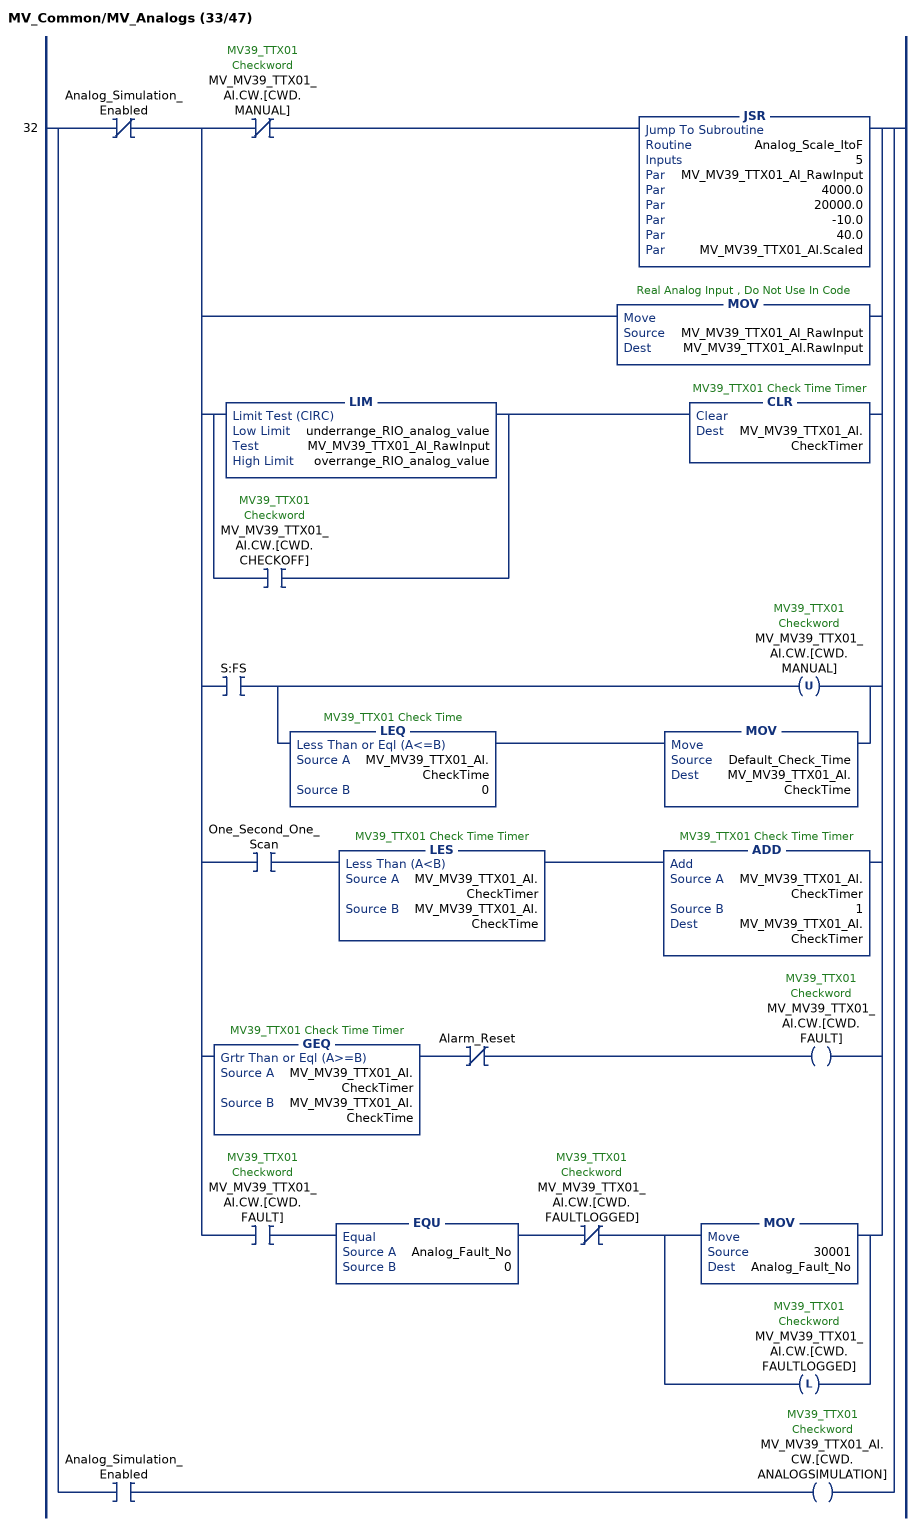
   32: [XIO(Analog_Simulation_Enabled) [XIO(MV_MV39_TTX01_AI.CW.[CWD.MANUAL]) JSR(Analog_Scale_ItoF,5,MV_MV39_TTX01_AI_RawInput,4000.0,20000.0,-10.0,40.0,MV_MV39_TTX01_AI.Scaled) ,MOV(MV_MV39_TTX01_AI_RawInput,MV_MV39_TTX01_AI.RawInput) ,[LIM(underrange_RIO_analog_value,MV_MV39_TTX01_AI_RawInput,overrange_RIO_analog_value) ,XIC(MV_MV39_TTX01_AI.CW.[CWD.CHECKOFF]) ] CLR(MV_MV39_TTX01_AI.CheckTimer) ,XIC(S:FS) [OTU(MV_MV39_TTX01_AI.CW.[CWD.MANUAL]) ,LEQ(MV_MV39_TTX01_AI.CheckTime,0) MOV(Default_Check_Time,MV_MV39_TTX01_AI.CheckTime) ] ,XIC(One_Second_One_Scan) LES(MV_MV39_TTX01_AI.CheckTimer,MV_MV39_TTX01_AI.CheckTime) ADD(MV_MV39_TTX01_AI.CheckTimer,1,MV_MV39_TTX01_AI.CheckTimer) ,GEQ(MV_MV39_TTX01_AI.CheckTimer,MV_MV39_TTX01_AI.CheckTime) XIO(Alarm_Reset) OTE(MV_MV39_TTX01_AI.CW.[CWD.FAULT]) ,XIC(MV_MV39_TTX01_AI.CW.[CWD.FAULT]) EQU(Analog_Fault_No,0) XIO(MV_MV39_TTX01_AI.CW.[CWD.FAULTLOGGED]) [MOV(30001,Analog_Fault_No) ,OTL(MV_MV39_TTX01_AI.CW.[CWD.FAULTLOGGED]) ] ] ,XIC(Analog_Simulation_Enabled) OTE(MV_MV39_TTX01_AI.CW.[CWD.ANALOGSIMULATION]) ];
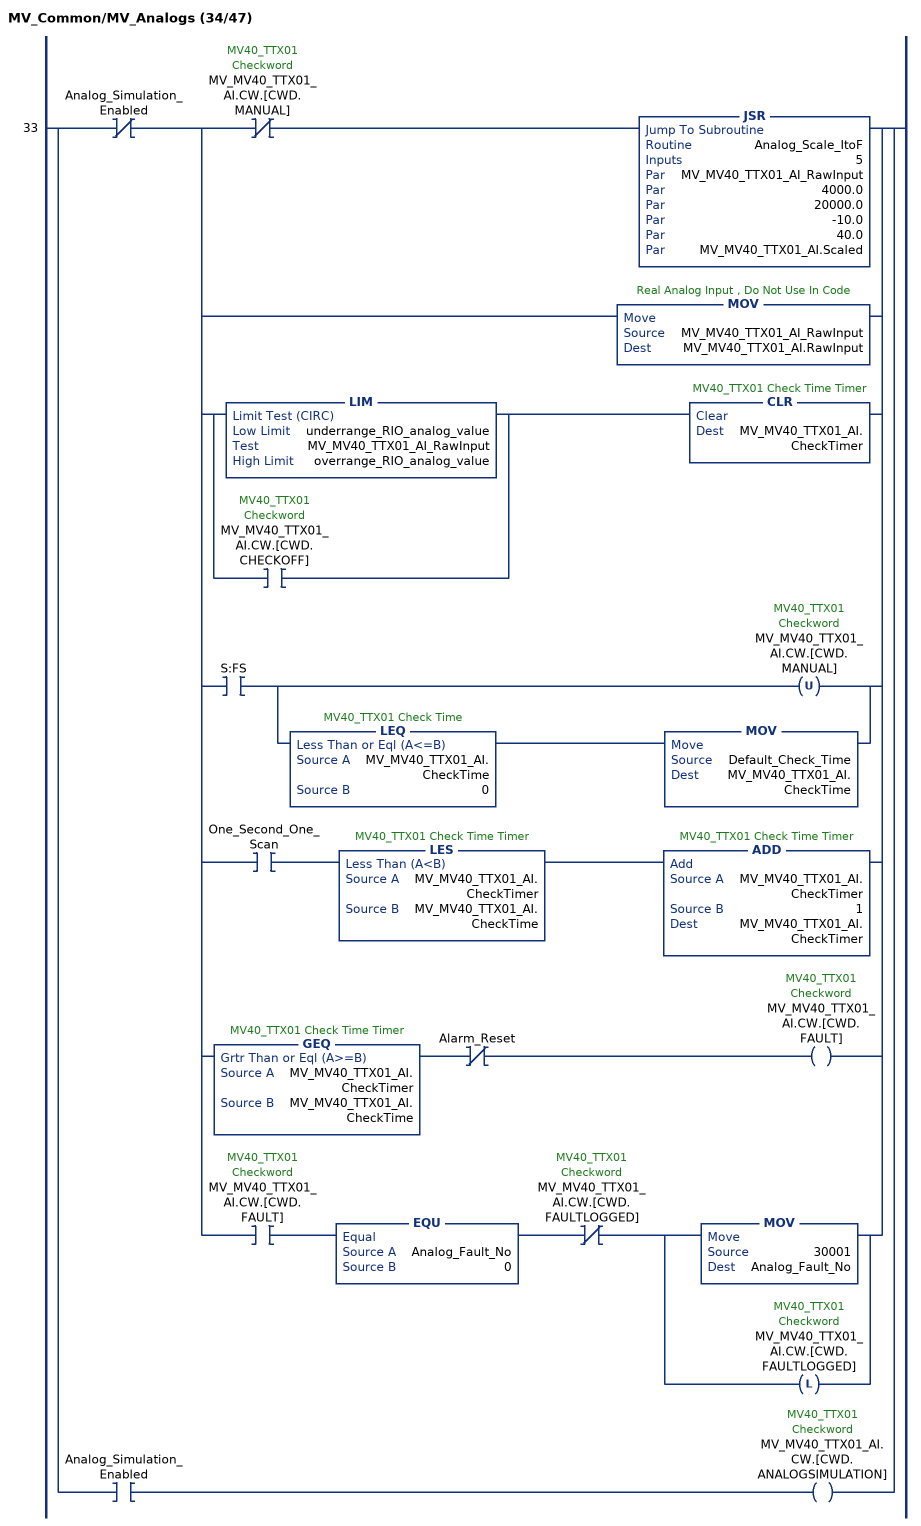
   33: [XIO(Analog_Simulation_Enabled) [XIO(MV_MV40_TTX01_AI.CW.[CWD.MANUAL]) JSR(Analog_Scale_ItoF,5,MV_MV40_TTX01_AI_RawInput,4000.0,20000.0,-10.0,40.0,MV_MV40_TTX01_AI.Scaled) ,MOV(MV_MV40_TTX01_AI_RawInput,MV_MV40_TTX01_AI.RawInput) ,[LIM(underrange_RIO_analog_value,MV_MV40_TTX01_AI_RawInput,overrange_RIO_analog_value) ,XIC(MV_MV40_TTX01_AI.CW.[CWD.CHECKOFF]) ] CLR(MV_MV40_TTX01_AI.CheckTimer) ,XIC(S:FS) [OTU(MV_MV40_TTX01_AI.CW.[CWD.MANUAL]) ,LEQ(MV_MV40_TTX01_AI.CheckTime,0) MOV(Default_Check_Time,MV_MV40_TTX01_AI.CheckTime) ] ,XIC(One_Second_One_Scan) LES(MV_MV40_TTX01_AI.CheckTimer,MV_MV40_TTX01_AI.CheckTime) ADD(MV_MV40_TTX01_AI.CheckTimer,1,MV_MV40_TTX01_AI.CheckTimer) ,GEQ(MV_MV40_TTX01_AI.CheckTimer,MV_MV40_TTX01_AI.CheckTime) XIO(Alarm_Reset) OTE(MV_MV40_TTX01_AI.CW.[CWD.FAULT]) ,XIC(MV_MV40_TTX01_AI.CW.[CWD.FAULT]) EQU(Analog_Fault_No,0) XIO(MV_MV40_TTX01_AI.CW.[CWD.FAULTLOGGED]) [MOV(30001,Analog_Fault_No) ,OTL(MV_MV40_TTX01_AI.CW.[CWD.FAULTLOGGED]) ] ] ,XIC(Analog_Simulation_Enabled) OTE(MV_MV40_TTX01_AI.CW.[CWD.ANALOGSIMULATION]) ];
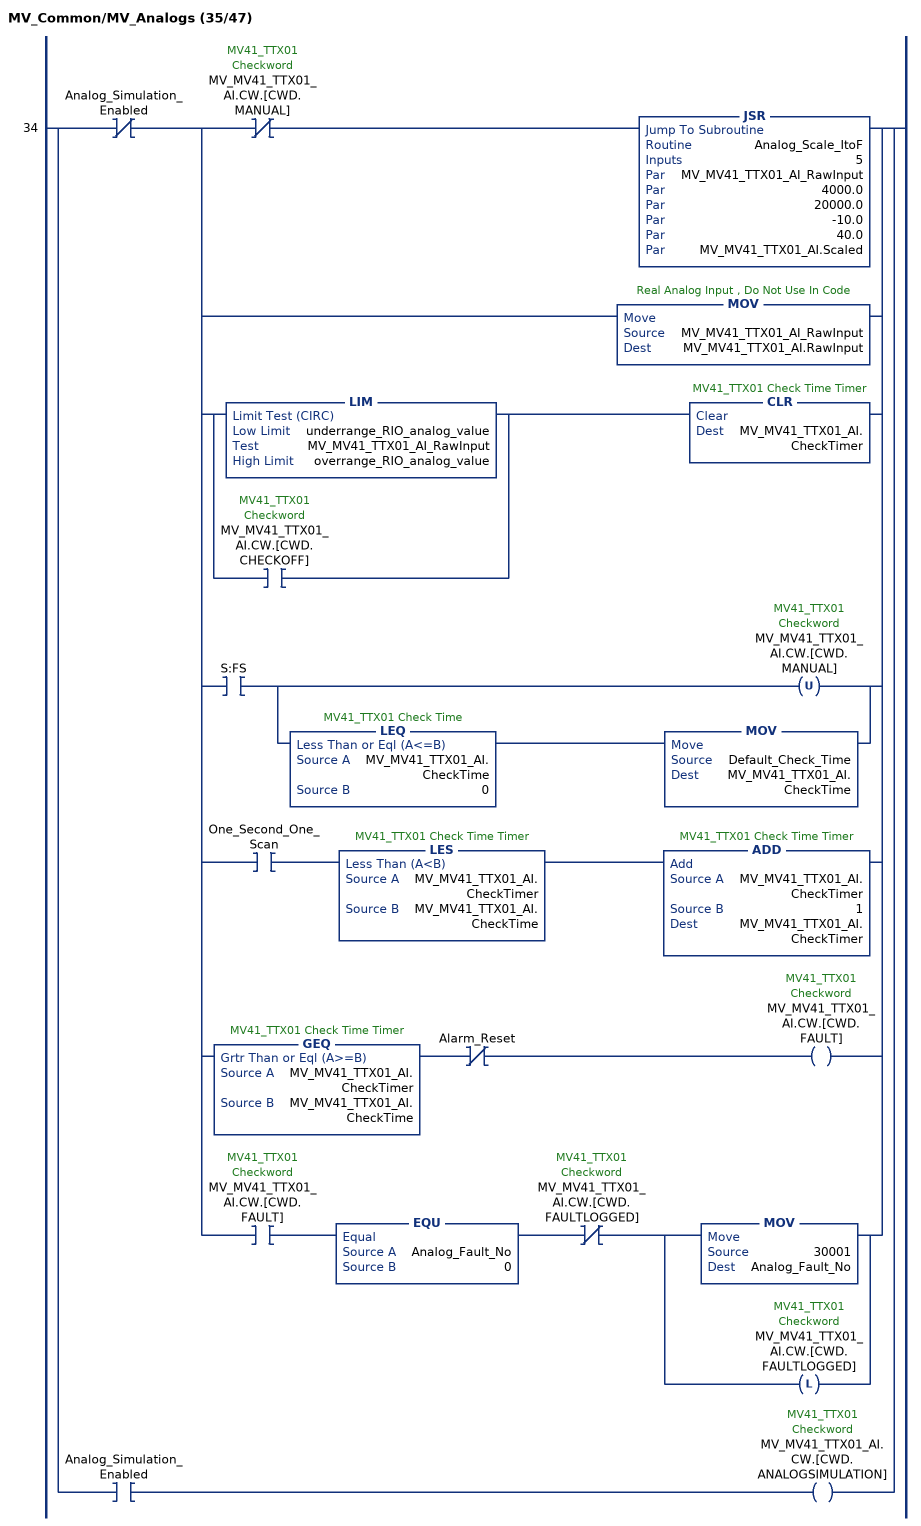
   34: [XIO(Analog_Simulation_Enabled) [XIO(MV_MV41_TTX01_AI.CW.[CWD.MANUAL]) JSR(Analog_Scale_ItoF,5,MV_MV41_TTX01_AI_RawInput,4000.0,20000.0,-10.0,40.0,MV_MV41_TTX01_AI.Scaled) ,MOV(MV_MV41_TTX01_AI_RawInput,MV_MV41_TTX01_AI.RawInput) ,[LIM(underrange_RIO_analog_value,MV_MV41_TTX01_AI_RawInput,overrange_RIO_analog_value) ,XIC(MV_MV41_TTX01_AI.CW.[CWD.CHECKOFF]) ] CLR(MV_MV41_TTX01_AI.CheckTimer) ,XIC(S:FS) [OTU(MV_MV41_TTX01_AI.CW.[CWD.MANUAL]) ,LEQ(MV_MV41_TTX01_AI.CheckTime,0) MOV(Default_Check_Time,MV_MV41_TTX01_AI.CheckTime) ] ,XIC(One_Second_One_Scan) LES(MV_MV41_TTX01_AI.CheckTimer,MV_MV41_TTX01_AI.CheckTime) ADD(MV_MV41_TTX01_AI.CheckTimer,1,MV_MV41_TTX01_AI.CheckTimer) ,GEQ(MV_MV41_TTX01_AI.CheckTimer,MV_MV41_TTX01_AI.CheckTime) XIO(Alarm_Reset) OTE(MV_MV41_TTX01_AI.CW.[CWD.FAULT]) ,XIC(MV_MV41_TTX01_AI.CW.[CWD.FAULT]) EQU(Analog_Fault_No,0) XIO(MV_MV41_TTX01_AI.CW.[CWD.FAULTLOGGED]) [MOV(30001,Analog_Fault_No) ,OTL(MV_MV41_TTX01_AI.CW.[CWD.FAULTLOGGED]) ] ] ,XIC(Analog_Simulation_Enabled) OTE(MV_MV41_TTX01_AI.CW.[CWD.ANALOGSIMULATION]) ];
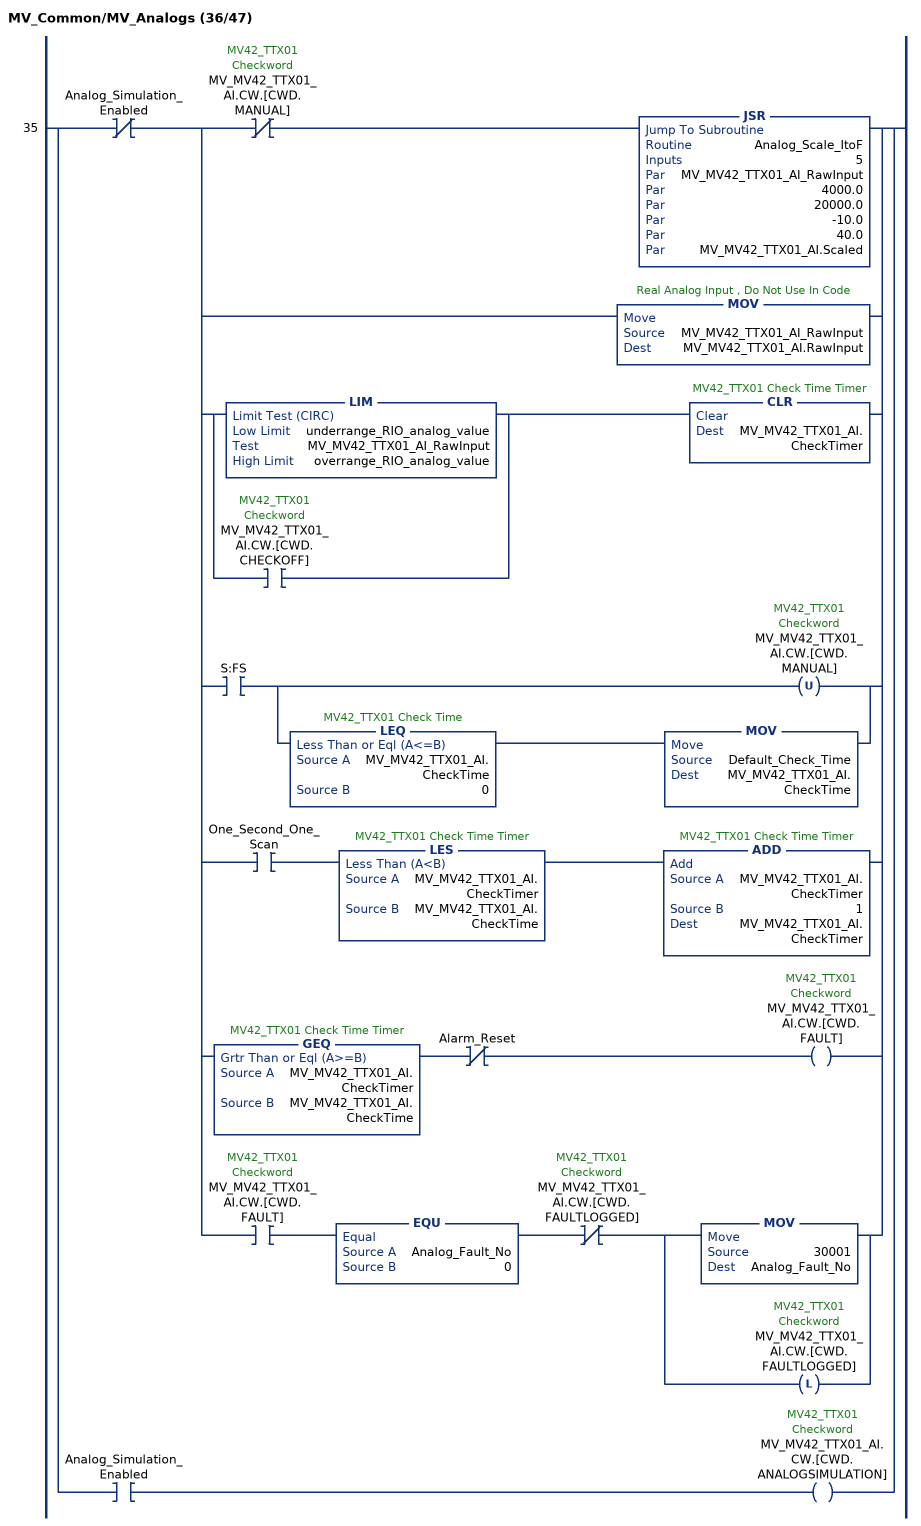
   35: [XIO(Analog_Simulation_Enabled) [XIO(MV_MV42_TTX01_AI.CW.[CWD.MANUAL]) JSR(Analog_Scale_ItoF,5,MV_MV42_TTX01_AI_RawInput,4000.0,20000.0,-10.0,40.0,MV_MV42_TTX01_AI.Scaled) ,MOV(MV_MV42_TTX01_AI_RawInput,MV_MV42_TTX01_AI.RawInput) ,[LIM(underrange_RIO_analog_value,MV_MV42_TTX01_AI_RawInput,overrange_RIO_analog_value) ,XIC(MV_MV42_TTX01_AI.CW.[CWD.CHECKOFF]) ] CLR(MV_MV42_TTX01_AI.CheckTimer) ,XIC(S:FS) [OTU(MV_MV42_TTX01_AI.CW.[CWD.MANUAL]) ,LEQ(MV_MV42_TTX01_AI.CheckTime,0) MOV(Default_Check_Time,MV_MV42_TTX01_AI.CheckTime) ] ,XIC(One_Second_One_Scan) LES(MV_MV42_TTX01_AI.CheckTimer,MV_MV42_TTX01_AI.CheckTime) ADD(MV_MV42_TTX01_AI.CheckTimer,1,MV_MV42_TTX01_AI.CheckTimer) ,GEQ(MV_MV42_TTX01_AI.CheckTimer,MV_MV42_TTX01_AI.CheckTime) XIO(Alarm_Reset) OTE(MV_MV42_TTX01_AI.CW.[CWD.FAULT]) ,XIC(MV_MV42_TTX01_AI.CW.[CWD.FAULT]) EQU(Analog_Fault_No,0) XIO(MV_MV42_TTX01_AI.CW.[CWD.FAULTLOGGED]) [MOV(30001,Analog_Fault_No) ,OTL(MV_MV42_TTX01_AI.CW.[CWD.FAULTLOGGED]) ] ] ,XIC(Analog_Simulation_Enabled) OTE(MV_MV42_TTX01_AI.CW.[CWD.ANALOGSIMULATION]) ];
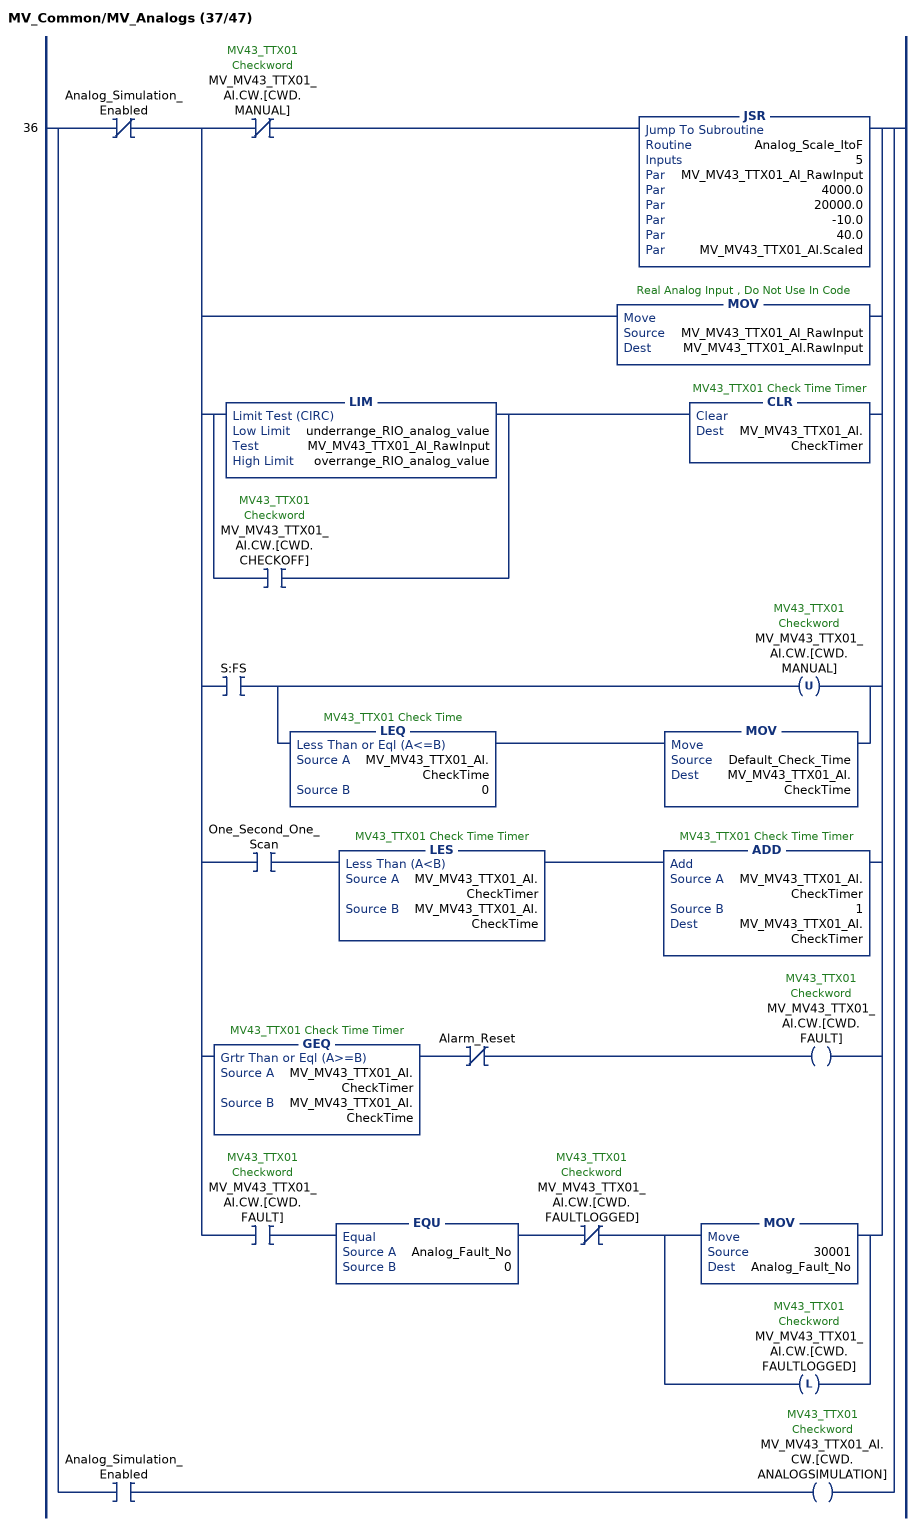
   36: [XIO(Analog_Simulation_Enabled) [XIO(MV_MV43_TTX01_AI.CW.[CWD.MANUAL]) JSR(Analog_Scale_ItoF,5,MV_MV43_TTX01_AI_RawInput,4000.0,20000.0,-10.0,40.0,MV_MV43_TTX01_AI.Scaled) ,MOV(MV_MV43_TTX01_AI_RawInput,MV_MV43_TTX01_AI.RawInput) ,[LIM(underrange_RIO_analog_value,MV_MV43_TTX01_AI_RawInput,overrange_RIO_analog_value) ,XIC(MV_MV43_TTX01_AI.CW.[CWD.CHECKOFF]) ] CLR(MV_MV43_TTX01_AI.CheckTimer) ,XIC(S:FS) [OTU(MV_MV43_TTX01_AI.CW.[CWD.MANUAL]) ,LEQ(MV_MV43_TTX01_AI.CheckTime,0) MOV(Default_Check_Time,MV_MV43_TTX01_AI.CheckTime) ] ,XIC(One_Second_One_Scan) LES(MV_MV43_TTX01_AI.CheckTimer,MV_MV43_TTX01_AI.CheckTime) ADD(MV_MV43_TTX01_AI.CheckTimer,1,MV_MV43_TTX01_AI.CheckTimer) ,GEQ(MV_MV43_TTX01_AI.CheckTimer,MV_MV43_TTX01_AI.CheckTime) XIO(Alarm_Reset) OTE(MV_MV43_TTX01_AI.CW.[CWD.FAULT]) ,XIC(MV_MV43_TTX01_AI.CW.[CWD.FAULT]) EQU(Analog_Fault_No,0) XIO(MV_MV43_TTX01_AI.CW.[CWD.FAULTLOGGED]) [MOV(30001,Analog_Fault_No) ,OTL(MV_MV43_TTX01_AI.CW.[CWD.FAULTLOGGED]) ] ] ,XIC(Analog_Simulation_Enabled) OTE(MV_MV43_TTX01_AI.CW.[CWD.ANALOGSIMULATION]) ];
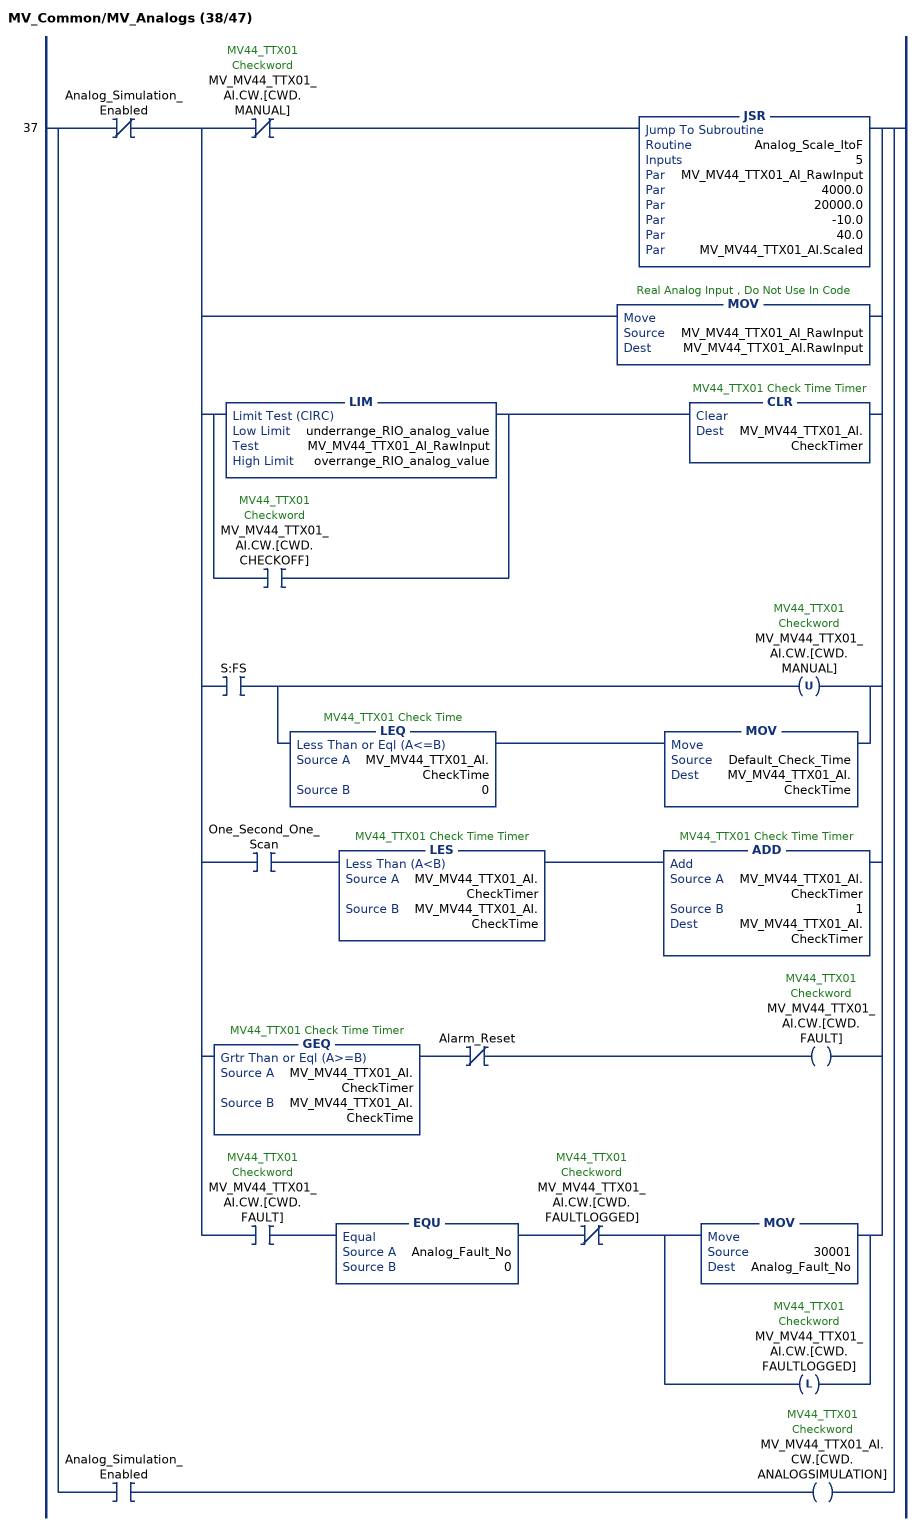
   37: [XIO(Analog_Simulation_Enabled) [XIO(MV_MV44_TTX01_AI.CW.[CWD.MANUAL]) JSR(Analog_Scale_ItoF,5,MV_MV44_TTX01_AI_RawInput,4000.0,20000.0,-10.0,40.0,MV_MV44_TTX01_AI.Scaled) ,MOV(MV_MV44_TTX01_AI_RawInput,MV_MV44_TTX01_AI.RawInput) ,[LIM(underrange_RIO_analog_value,MV_MV44_TTX01_AI_RawInput,overrange_RIO_analog_value) ,XIC(MV_MV44_TTX01_AI.CW.[CWD.CHECKOFF]) ] CLR(MV_MV44_TTX01_AI.CheckTimer) ,XIC(S:FS) [OTU(MV_MV44_TTX01_AI.CW.[CWD.MANUAL]) ,LEQ(MV_MV44_TTX01_AI.CheckTime,0) MOV(Default_Check_Time,MV_MV44_TTX01_AI.CheckTime) ] ,XIC(One_Second_One_Scan) LES(MV_MV44_TTX01_AI.CheckTimer,MV_MV44_TTX01_AI.CheckTime) ADD(MV_MV44_TTX01_AI.CheckTimer,1,MV_MV44_TTX01_AI.CheckTimer) ,GEQ(MV_MV44_TTX01_AI.CheckTimer,MV_MV44_TTX01_AI.CheckTime) XIO(Alarm_Reset) OTE(MV_MV44_TTX01_AI.CW.[CWD.FAULT]) ,XIC(MV_MV44_TTX01_AI.CW.[CWD.FAULT]) EQU(Analog_Fault_No,0) XIO(MV_MV44_TTX01_AI.CW.[CWD.FAULTLOGGED]) [MOV(30001,Analog_Fault_No) ,OTL(MV_MV44_TTX01_AI.CW.[CWD.FAULTLOGGED]) ] ] ,XIC(Analog_Simulation_Enabled) OTE(MV_MV44_TTX01_AI.CW.[CWD.ANALOGSIMULATION]) ];
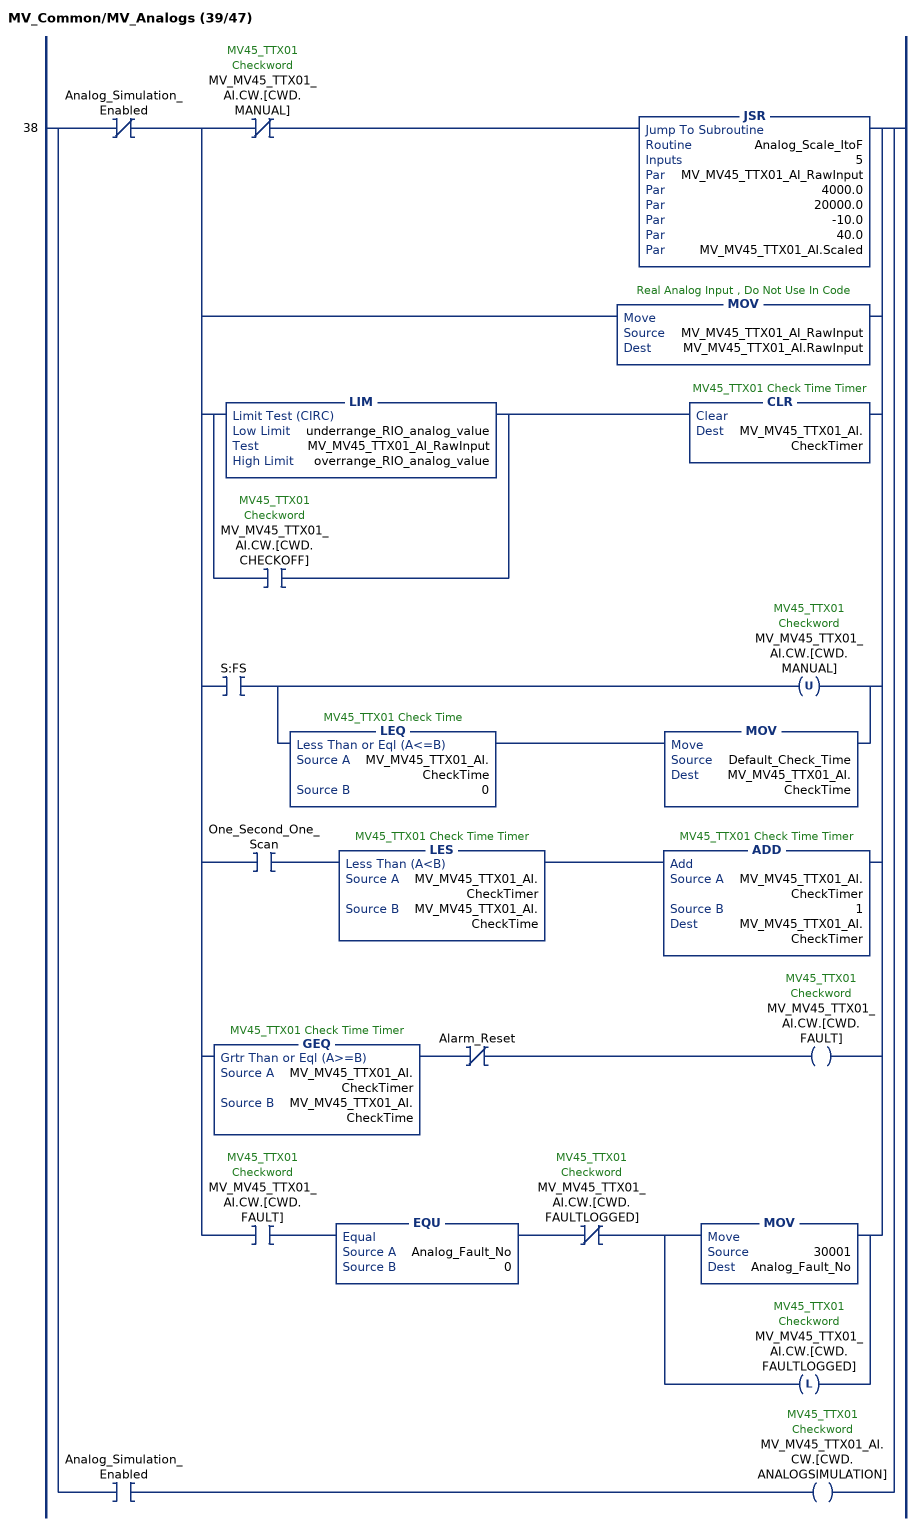
   38: [XIO(Analog_Simulation_Enabled) [XIO(MV_MV45_TTX01_AI.CW.[CWD.MANUAL]) JSR(Analog_Scale_ItoF,5,MV_MV45_TTX01_AI_RawInput,4000.0,20000.0,-10.0,40.0,MV_MV45_TTX01_AI.Scaled) ,MOV(MV_MV45_TTX01_AI_RawInput,MV_MV45_TTX01_AI.RawInput) ,[LIM(underrange_RIO_analog_value,MV_MV45_TTX01_AI_RawInput,overrange_RIO_analog_value) ,XIC(MV_MV45_TTX01_AI.CW.[CWD.CHECKOFF]) ] CLR(MV_MV45_TTX01_AI.CheckTimer) ,XIC(S:FS) [OTU(MV_MV45_TTX01_AI.CW.[CWD.MANUAL]) ,LEQ(MV_MV45_TTX01_AI.CheckTime,0) MOV(Default_Check_Time,MV_MV45_TTX01_AI.CheckTime) ] ,XIC(One_Second_One_Scan) LES(MV_MV45_TTX01_AI.CheckTimer,MV_MV45_TTX01_AI.CheckTime) ADD(MV_MV45_TTX01_AI.CheckTimer,1,MV_MV45_TTX01_AI.CheckTimer) ,GEQ(MV_MV45_TTX01_AI.CheckTimer,MV_MV45_TTX01_AI.CheckTime) XIO(Alarm_Reset) OTE(MV_MV45_TTX01_AI.CW.[CWD.FAULT]) ,XIC(MV_MV45_TTX01_AI.CW.[CWD.FAULT]) EQU(Analog_Fault_No,0) XIO(MV_MV45_TTX01_AI.CW.[CWD.FAULTLOGGED]) [MOV(30001,Analog_Fault_No) ,OTL(MV_MV45_TTX01_AI.CW.[CWD.FAULTLOGGED]) ] ] ,XIC(Analog_Simulation_Enabled) OTE(MV_MV45_TTX01_AI.CW.[CWD.ANALOGSIMULATION]) ];
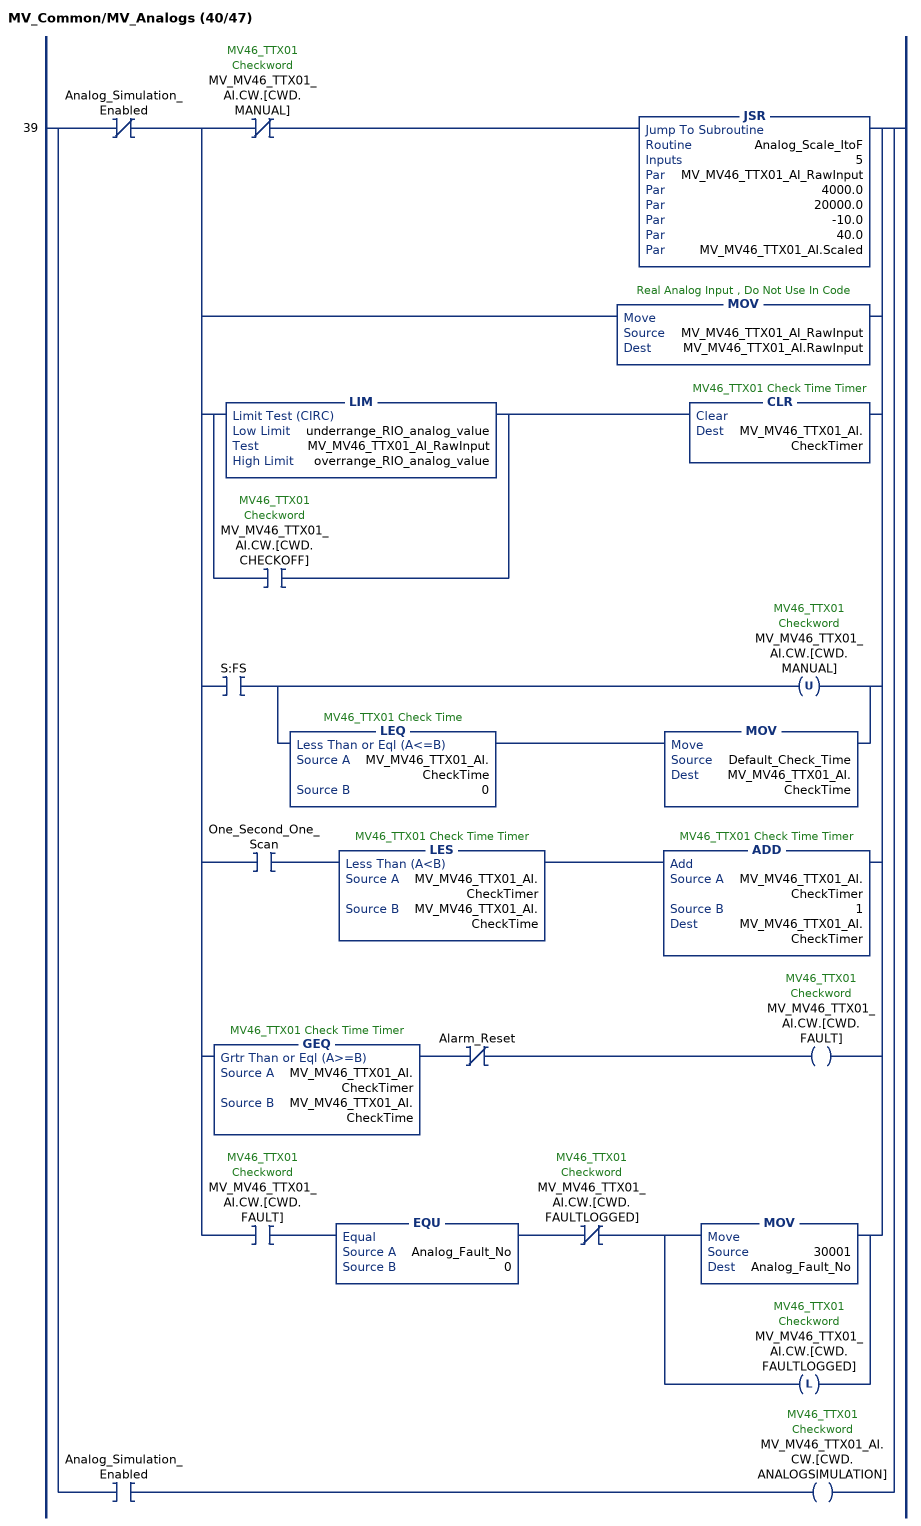
   39: [XIO(Analog_Simulation_Enabled) [XIO(MV_MV46_TTX01_AI.CW.[CWD.MANUAL]) JSR(Analog_Scale_ItoF,5,MV_MV46_TTX01_AI_RawInput,4000.0,20000.0,-10.0,40.0,MV_MV46_TTX01_AI.Scaled) ,MOV(MV_MV46_TTX01_AI_RawInput,MV_MV46_TTX01_AI.RawInput) ,[LIM(underrange_RIO_analog_value,MV_MV46_TTX01_AI_RawInput,overrange_RIO_analog_value) ,XIC(MV_MV46_TTX01_AI.CW.[CWD.CHECKOFF]) ] CLR(MV_MV46_TTX01_AI.CheckTimer) ,XIC(S:FS) [OTU(MV_MV46_TTX01_AI.CW.[CWD.MANUAL]) ,LEQ(MV_MV46_TTX01_AI.CheckTime,0) MOV(Default_Check_Time,MV_MV46_TTX01_AI.CheckTime) ] ,XIC(One_Second_One_Scan) LES(MV_MV46_TTX01_AI.CheckTimer,MV_MV46_TTX01_AI.CheckTime) ADD(MV_MV46_TTX01_AI.CheckTimer,1,MV_MV46_TTX01_AI.CheckTimer) ,GEQ(MV_MV46_TTX01_AI.CheckTimer,MV_MV46_TTX01_AI.CheckTime) XIO(Alarm_Reset) OTE(MV_MV46_TTX01_AI.CW.[CWD.FAULT]) ,XIC(MV_MV46_TTX01_AI.CW.[CWD.FAULT]) EQU(Analog_Fault_No,0) XIO(MV_MV46_TTX01_AI.CW.[CWD.FAULTLOGGED]) [MOV(30001,Analog_Fault_No) ,OTL(MV_MV46_TTX01_AI.CW.[CWD.FAULTLOGGED]) ] ] ,XIC(Analog_Simulation_Enabled) OTE(MV_MV46_TTX01_AI.CW.[CWD.ANALOGSIMULATION]) ];
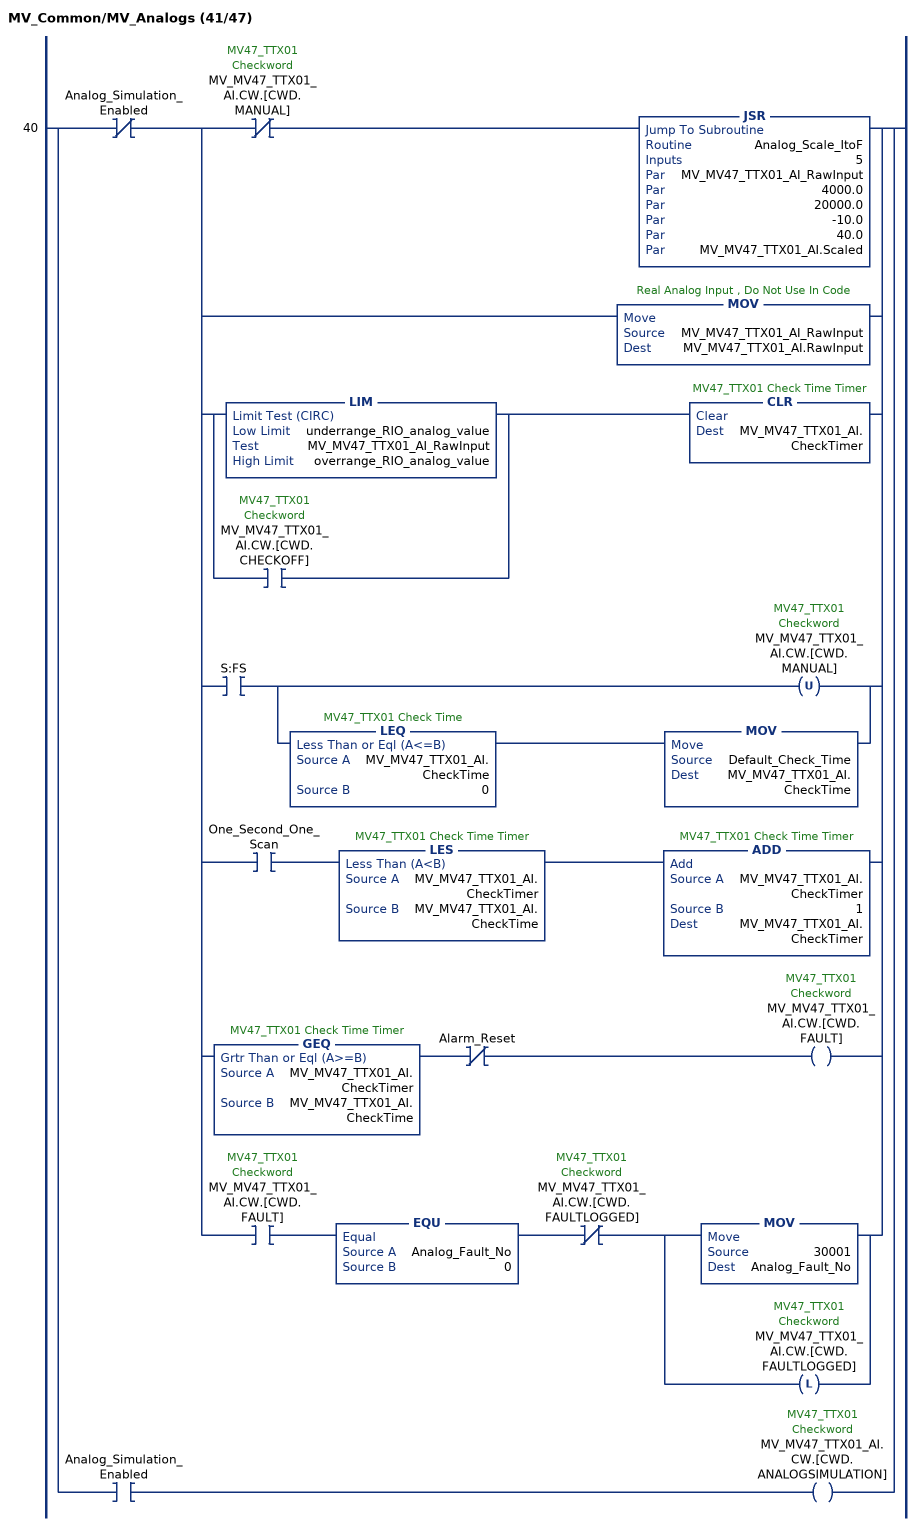
   40: [XIO(Analog_Simulation_Enabled) [XIO(MV_MV47_TTX01_AI.CW.[CWD.MANUAL]) JSR(Analog_Scale_ItoF,5,MV_MV47_TTX01_AI_RawInput,4000.0,20000.0,-10.0,40.0,MV_MV47_TTX01_AI.Scaled) ,MOV(MV_MV47_TTX01_AI_RawInput,MV_MV47_TTX01_AI.RawInput) ,[LIM(underrange_RIO_analog_value,MV_MV47_TTX01_AI_RawInput,overrange_RIO_analog_value) ,XIC(MV_MV47_TTX01_AI.CW.[CWD.CHECKOFF]) ] CLR(MV_MV47_TTX01_AI.CheckTimer) ,XIC(S:FS) [OTU(MV_MV47_TTX01_AI.CW.[CWD.MANUAL]) ,LEQ(MV_MV47_TTX01_AI.CheckTime,0) MOV(Default_Check_Time,MV_MV47_TTX01_AI.CheckTime) ] ,XIC(One_Second_One_Scan) LES(MV_MV47_TTX01_AI.CheckTimer,MV_MV47_TTX01_AI.CheckTime) ADD(MV_MV47_TTX01_AI.CheckTimer,1,MV_MV47_TTX01_AI.CheckTimer) ,GEQ(MV_MV47_TTX01_AI.CheckTimer,MV_MV47_TTX01_AI.CheckTime) XIO(Alarm_Reset) OTE(MV_MV47_TTX01_AI.CW.[CWD.FAULT]) ,XIC(MV_MV47_TTX01_AI.CW.[CWD.FAULT]) EQU(Analog_Fault_No,0) XIO(MV_MV47_TTX01_AI.CW.[CWD.FAULTLOGGED]) [MOV(30001,Analog_Fault_No) ,OTL(MV_MV47_TTX01_AI.CW.[CWD.FAULTLOGGED]) ] ] ,XIC(Analog_Simulation_Enabled) OTE(MV_MV47_TTX01_AI.CW.[CWD.ANALOGSIMULATION]) ];
